(* Logix 5000 project; controller OWF Emulate 5570 rev 30.12; software revision 30.00 *)

TASK MainTask (periodic, rate 1000 ms, priority 1, watchdog 5000 ms) : MainProgram

MODULES
   Local : Emulate 5570 (ICP 2, rev 30.12)
       : vendor 1 type 0 code 15 (ICP 0, rev 1.1, Output RPI 50 ms)
END_MODULES

TYPE UDT_BA :
STRUCT
   AL : BOOL[128];
END_STRUCT
END_TYPE

PROGRAM MainProgram   (* main routine MainRoutine *)
VAR
   OWF_Add_c : DINT;
   OWF_bit : DINT;
   OWF_blk : DINT;
   OWF_i : DINT;
   OWF_Input : DINT[16];
   OWF_InputLen : DINT;
   OWF_InputMaxInd : DINT;
   OWF_j : DINT;
   OWF_Key : DINT[512,17];
   OWF_Result : DINT[17];
   OWF_Ver : DINT;
   SCAN_CYCLE_TIME : DINT;
END_VAR

ROUTINE Application   (* structured text *)
   //Description: initialize the variables.
   
   if S:FS then  (* this is the first, normal scan of the routines in the current program, initialize the program.*)
   	OWF_Ver:=2;  //OWF_Ver means that the version of OWF: 256-256 bits, 384-384 bits, and 512-512 bits. The first number is length of input, the last number is length of output.
                    //If OWF_Ver means that the version of Hash, then three versions are: 256-128 bits, 384-160 bits and 512-256 bits.
   	If OWF_Ver=0 then
   		OWF_InputLen:=255;  //bits of input.
   		OWF_InputMaxInd:=8;  //maximum index for dints which store the bits of input.
   		for OWF_i:=0 to OWF_InputMaxInd-1 by 1 Do
   			//OWF_Input[OWF_i]:= 65535;   //Half of the selection factors are 1.
   			OWF_Input[OWF_i]:= -1;    //All the selection factors are 1.
   		end_for;
   	end_if;
   
   
   	If OWF_Ver=1 then
   		OWF_InputLen:= 383;
   		OWF_InputMaxInd:=12;  //maximum index for array.
   		for OWF_i:=0 to OWF_InputMaxInd-1 by 1 Do
   			//OWF_Input[OWF_i]:= 65535;     //Half of the selection factors are 1.
   			OWF_Input[OWF_i]:= -1;   //All the selection factors are 1.
   		end_for;
   	end_if;
   
   
   	If OWF_Ver=2 then
   		OWF_InputLen:= 511;
   		OWF_InputMaxInd:=16;  //maximum index for array.
   		for OWF_i:=0 to OWF_InputMaxInd-1 by 1 Do
   			//OWF_Input[OWF_i]:= 65535;     //Half of the selection factors are 1.
   			OWF_Input[OWF_i]:= -1;   //All the selection factors are 1.
   		end_for;
   	end_if;
   
   end_if;
   
   
   
   
   
END_ROUTINE

ROUTINE MainRoutine   (* ladder *)
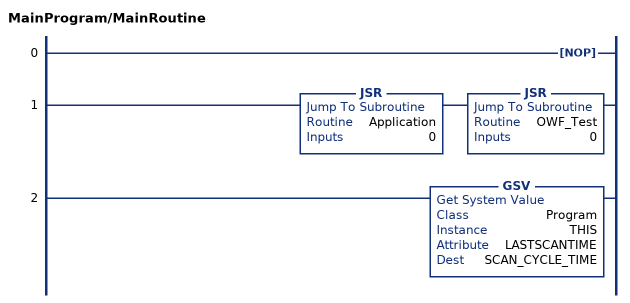
   0: NOP();
   1: JSR(Application,0)JSR(OWF_Test,0);
   2: GSV(Program,THIS,LASTSCANTIME,SCAN_CYCLE_TIME);
END_ROUTINE

ROUTINE Original_OWF   (* structured text *)
   
   //implement One Way Function (OWF) based on subset Sum.
   //input: choice factor OWF_Input[], array OWF_Key[][].
   //output: OWF_Result[]
   
   (*
   	for OWF_i:=0 to OWF_InputMaxInd by 1 Do
   		OWF_Result[OWF_i]:= 0;  //Initialize the OWF_Result[].
   	end_for;
   *)
   
   
   OWF_bit:=0;   // bit index
   OWF_blk:=0;   // block index
   
   JSR(OWF_Init);
   
   	//compute subset sum.
   	for OWF_i:=0 to OWF_InputLen by 1 do
   		If OWF_bit = 32 then
   			OWF_bit:=0;
   			OWF_blk:=OWF_blk+1;
   		end_if;
   		OWF_Add_c:=0;
   		if OWF_Input[OWF_blk].[OWF_bit] then
   			for OWF_j:=0 to OWF_InputMaxInd-1 by 1 Do
   				OWF_Result[OWF_j]:=OWF_Result[OWF_j] + OWF_Key[OWF_i,OWF_j] + OWF_Add_c;    //compute the result of subset sum.
   				OWF_Add_c.0:= OWF_Result[OWF_j].31;
   				OWF_Result[OWF_j].31:=0;
   			end_for;
   			OWF_Result[OWF_j]:=OWF_Result[OWF_j] + OWF_Key[OWF_i,OWF_j] + OWF_Add_c;
   		end_if;
   		OWF_bit:=OWF_bit + 1;
   	end_for;
   
   If OWF_Ver=0 Then
   	OWF_Result[OWF_InputMaxInd]:=OWF_Result[OWF_InputMaxInd] and 16#FF; //clear high bit
   End_If;
   
   If OWF_Ver=1 Then
   	OWF_Result[OWF_InputMaxInd]:=OWF_Result[OWF_InputMaxInd] and 16#FFF; //clear high bit
   End_If;
   
   If OWF_Ver = 2 Then
   	OWF_Result[OWF_InputMaxInd]:=OWF_Result[OWF_InputMaxInd] and 16#FFFF; //clear high bit
   End_If;
END_ROUTINE

ROUTINE OWF_Init   (* structured text *)
   If OWF_Ver >= 0 Then
   	OWF_Key[0,0]:=1227121054;
   	OWF_Key[0,1]:=202649963;
   	OWF_Key[0,2]:=1031163235;
   	OWF_Key[0,3]:=558332383;
   	OWF_Key[0,4]:=758449748;
   	OWF_Key[0,5]:=439100062;
   	OWF_Key[0,6]:=1763017217;
   	OWF_Key[0,7]:=741113131;
   	OWF_Key[0,8]:=1652892808;
   	OWF_Key[1,0]:=1354606577;
   	OWF_Key[1,1]:=1085346626;
   	OWF_Key[1,2]:=1684734244;
   	OWF_Key[1,3]:=1525280682;
   	OWF_Key[1,4]:=581896247;
   	OWF_Key[1,5]:=1418880834;
   	OWF_Key[1,6]:=1348359995;
   	OWF_Key[1,7]:=1446005479;
   	OWF_Key[1,8]:=332839494;
   	OWF_Key[2,0]:=2095017041;
   	OWF_Key[2,1]:=1217317816;
   	OWF_Key[2,2]:=648181522;
   	OWF_Key[2,3]:=178964298;
   	OWF_Key[2,4]:=463461758;
   	OWF_Key[2,5]:=346394231;
   	OWF_Key[2,6]:=1486999699;
   	OWF_Key[2,7]:=1770617031;
   	OWF_Key[2,8]:=362139479;
   	OWF_Key[3,0]:=256347809;
   	OWF_Key[3,1]:=1312207174;
   	OWF_Key[3,2]:=843085075;
   	OWF_Key[3,3]:=1139982972;
   	OWF_Key[3,4]:=662387156;
   	OWF_Key[3,5]:=1025052915;
   	OWF_Key[3,6]:=1908648583;
   	OWF_Key[3,7]:=1963224943;
   	OWF_Key[3,8]:=1427256681;
   	OWF_Key[4,0]:=1972101745;
   	OWF_Key[4,1]:=1002975333;
   	OWF_Key[4,2]:=1871427740;
   	OWF_Key[4,3]:=1318551426;
   	OWF_Key[4,4]:=1364597906;
   	OWF_Key[4,5]:=1294123204;
   	OWF_Key[4,6]:=2125414218;
   	OWF_Key[4,7]:=1926341024;
   	OWF_Key[4,8]:=460259043;
   	OWF_Key[5,0]:=1524399156;
   	OWF_Key[5,1]:=2011514619;
   	OWF_Key[5,2]:=2069350563;
   	OWF_Key[5,3]:=279858814;
   	OWF_Key[5,4]:=810485067;
   	OWF_Key[5,5]:=73617388;
   	OWF_Key[5,6]:=687884215;
   	OWF_Key[5,7]:=1340310677;
   	OWF_Key[5,8]:=431345285;
   	OWF_Key[6,0]:=1066476071;
   	OWF_Key[6,1]:=550806088;
   	OWF_Key[6,2]:=756174308;
   	OWF_Key[6,3]:=574071763;
   	OWF_Key[6,4]:=409094206;
   	OWF_Key[6,5]:=1665642823;
   	OWF_Key[6,6]:=1813040245;
   	OWF_Key[6,7]:=215573695;
   	OWF_Key[6,8]:=525097691;
   	OWF_Key[7,0]:=1934399231;
   	OWF_Key[7,1]:=1553053230;
   	OWF_Key[7,2]:=144946822;
   	OWF_Key[7,3]:=2140599730;
   	OWF_Key[7,4]:=1889193085;
   	OWF_Key[7,5]:=2054644962;
   	OWF_Key[7,6]:=826013297;
   	OWF_Key[7,7]:=556817065;
   	OWF_Key[7,8]:=33718400;
   	OWF_Key[8,0]:=899651387;
   	OWF_Key[8,1]:=1251867014;
   	OWF_Key[8,2]:=959094800;
   	OWF_Key[8,3]:=194574689;
   	OWF_Key[8,4]:=1642465144;
   	OWF_Key[8,5]:=1096334976;
   	OWF_Key[8,6]:=931056050;
   	OWF_Key[8,7]:=405780298;
   	OWF_Key[8,8]:=1355752490;
   	OWF_Key[9,0]:=1528579024;
   	OWF_Key[9,1]:=1525333419;
   	OWF_Key[9,2]:=1348534735;
   	OWF_Key[9,3]:=111603084;
   	OWF_Key[9,4]:=1832745100;
   	OWF_Key[9,5]:=642195240;
   	OWF_Key[9,6]:=966181946;
   	OWF_Key[9,7]:=880029259;
   	OWF_Key[9,8]:=1162642342;
   	OWF_Key[10,0]:=359569674;
   	OWF_Key[10,1]:=1980700574;
   	OWF_Key[10,2]:=1293914236;
   	OWF_Key[10,3]:=954723255;
   	OWF_Key[10,4]:=1377909373;
   	OWF_Key[10,5]:=223244700;
   	OWF_Key[10,6]:=1984808221;
   	OWF_Key[10,7]:=1498924409;
   	OWF_Key[10,8]:=29167191;
   	OWF_Key[11,0]:=623116396;
   	OWF_Key[11,1]:=256225512;
   	OWF_Key[11,2]:=1328608936;
   	OWF_Key[11,3]:=725706243;
   	OWF_Key[11,4]:=791017754;
   	OWF_Key[11,5]:=1341758946;
   	OWF_Key[11,6]:=1113167772;
   	OWF_Key[11,7]:=639937104;
   	OWF_Key[11,8]:=436330960;
   	OWF_Key[12,0]:=1329424307;
   	OWF_Key[12,1]:=101924380;
   	OWF_Key[12,2]:=1635207076;
   	OWF_Key[12,3]:=1264309098;
   	OWF_Key[12,4]:=1613321141;
   	OWF_Key[12,5]:=1843793655;
   	OWF_Key[12,6]:=1519128380;
   	OWF_Key[12,7]:=1637695475;
   	OWF_Key[12,8]:=1595160782;
   	OWF_Key[13,0]:=475438733;
   	OWF_Key[13,1]:=914493831;
   	OWF_Key[13,2]:=239185193;
   	OWF_Key[13,3]:=7070920;
   	OWF_Key[13,4]:=1909091689;
   	OWF_Key[13,5]:=818931882;
   	OWF_Key[13,6]:=167044628;
   	OWF_Key[13,7]:=1264941904;
   	OWF_Key[13,8]:=949875305;
   	OWF_Key[14,0]:=1115356298;
   	OWF_Key[14,1]:=338497818;
   	OWF_Key[14,2]:=180024891;
   	OWF_Key[14,3]:=844456349;
   	OWF_Key[14,4]:=1506829383;
   	OWF_Key[14,5]:=94052327;
   	OWF_Key[14,6]:=1993991460;
   	OWF_Key[14,7]:=23038222;
   	OWF_Key[14,8]:=87146691;
   	OWF_Key[15,0]:=326487164;
   	OWF_Key[15,1]:=516484364;
   	OWF_Key[15,2]:=1296941749;
   	OWF_Key[15,3]:=811092697;
   	OWF_Key[15,4]:=538927605;
   	OWF_Key[15,5]:=659414599;
   	OWF_Key[15,6]:=759387250;
   	OWF_Key[15,7]:=589772068;
   	OWF_Key[15,8]:=514624038;
   	OWF_Key[16,0]:=1091875462;
   	OWF_Key[16,1]:=461268148;
   	OWF_Key[16,2]:=1603288957;
   	OWF_Key[16,3]:=626416433;
   	OWF_Key[16,4]:=654301897;
   	OWF_Key[16,5]:=1861165437;
   	OWF_Key[16,6]:=710648683;
   	OWF_Key[16,7]:=706991177;
   	OWF_Key[16,8]:=2023521577;
   	OWF_Key[17,0]:=1533914360;
   	OWF_Key[17,1]:=2033382504;
   	OWF_Key[17,2]:=1913483458;
   	OWF_Key[17,3]:=1068320764;
   	OWF_Key[17,4]:=1873217994;
   	OWF_Key[17,5]:=462057421;
   	OWF_Key[17,6]:=434206996;
   	OWF_Key[17,7]:=967662215;
   	OWF_Key[17,8]:=1066362328;
   	OWF_Key[18,0]:=1233616361;
   	OWF_Key[18,1]:=1376108010;
   	OWF_Key[18,2]:=151681671;
   	OWF_Key[18,3]:=1118724616;
   	OWF_Key[18,4]:=870582805;
   	OWF_Key[18,5]:=838422454;
   	OWF_Key[18,6]:=958525863;
   	OWF_Key[18,7]:=884926077;
   	OWF_Key[18,8]:=1110871443;
   	OWF_Key[19,0]:=1105934356;
   	OWF_Key[19,1]:=664442467;
   	OWF_Key[19,2]:=903233013;
   	OWF_Key[19,3]:=987099294;
   	OWF_Key[19,4]:=737604300;
   	OWF_Key[19,5]:=1759631091;
   	OWF_Key[19,6]:=1580233890;
   	OWF_Key[19,7]:=1669577827;
   	OWF_Key[19,8]:=91657386;
   	OWF_Key[20,0]:=360120849;
   	OWF_Key[20,1]:=1832314473;
   	OWF_Key[20,2]:=2086185527;
   	OWF_Key[20,3]:=1076864314;
   	OWF_Key[20,4]:=1498905358;
   	OWF_Key[20,5]:=900988985;
   	OWF_Key[20,6]:=1478986721;
   	OWF_Key[20,7]:=1681057774;
   	OWF_Key[20,8]:=562389748;
   	OWF_Key[21,0]:=368575225;
   	OWF_Key[21,1]:=2040057957;
   	OWF_Key[21,2]:=1772443406;
   	OWF_Key[21,3]:=358038348;
   	OWF_Key[21,4]:=1880468616;
   	OWF_Key[21,5]:=1275762442;
   	OWF_Key[21,6]:=240738790;
   	OWF_Key[21,7]:=1742748974;
   	OWF_Key[21,8]:=1288995313;
   	OWF_Key[22,0]:=2102585710;
   	OWF_Key[22,1]:=1254850839;
   	OWF_Key[22,2]:=1750685415;
   	OWF_Key[22,3]:=407311703;
   	OWF_Key[22,4]:=1927455536;
   	OWF_Key[22,5]:=734780728;
   	OWF_Key[22,6]:=1963803180;
   	OWF_Key[22,7]:=24276587;
   	OWF_Key[22,8]:=305836334;
   	OWF_Key[23,0]:=1060880211;
   	OWF_Key[23,1]:=321236053;
   	OWF_Key[23,2]:=1978313959;
   	OWF_Key[23,3]:=280999634;
   	OWF_Key[23,4]:=811422929;
   	OWF_Key[23,5]:=1151495141;
   	OWF_Key[23,6]:=684998164;
   	OWF_Key[23,7]:=1774640068;
   	OWF_Key[23,8]:=1081430675;
   	OWF_Key[24,0]:=1100474918;
   	OWF_Key[24,1]:=604700422;
   	OWF_Key[24,2]:=1689758319;
   	OWF_Key[24,3]:=215570041;
   	OWF_Key[24,4]:=1701438018;
   	OWF_Key[24,5]:=1754755041;
   	OWF_Key[24,6]:=7425442;
   	OWF_Key[24,7]:=918208170;
   	OWF_Key[24,8]:=1719377360;
   	OWF_Key[25,0]:=1547355790;
   	OWF_Key[25,1]:=1403608030;
   	OWF_Key[25,2]:=1499880269;
   	OWF_Key[25,3]:=317100104;
   	OWF_Key[25,4]:=1905628845;
   	OWF_Key[25,5]:=1066486402;
   	OWF_Key[25,6]:=756239231;
   	OWF_Key[25,7]:=459531339;
   	OWF_Key[25,8]:=1346452392;
   	OWF_Key[26,0]:=168483711;
   	OWF_Key[26,1]:=1800574949;
   	OWF_Key[26,2]:=1200797705;
   	OWF_Key[26,3]:=14565181;
   	OWF_Key[26,4]:=228173521;
   	OWF_Key[26,5]:=1764496443;
   	OWF_Key[26,6]:=504637489;
   	OWF_Key[26,7]:=1780840621;
   	OWF_Key[26,8]:=1379082303;
   	OWF_Key[27,0]:=54123181;
   	OWF_Key[27,1]:=622944351;
   	OWF_Key[27,2]:=2100500392;
   	OWF_Key[27,3]:=1775742704;
   	OWF_Key[27,4]:=143633756;
   	OWF_Key[27,5]:=1536231566;
   	OWF_Key[27,6]:=1440183257;
   	OWF_Key[27,7]:=2114239512;
   	OWF_Key[27,8]:=53396177;
   	OWF_Key[28,0]:=2134211248;
   	OWF_Key[28,1]:=1985332782;
   	OWF_Key[28,2]:=660997500;
   	OWF_Key[28,3]:=1607311701;
   	OWF_Key[28,4]:=1401991464;
   	OWF_Key[28,5]:=891355717;
   	OWF_Key[28,6]:=1475041716;
   	OWF_Key[28,7]:=258011330;
   	OWF_Key[28,8]:=2098653906;
   	OWF_Key[29,0]:=1790937980;
   	OWF_Key[29,1]:=592851196;
   	OWF_Key[29,2]:=1910540181;
   	OWF_Key[29,3]:=664243004;
   	OWF_Key[29,4]:=360474841;
   	OWF_Key[29,5]:=1110300911;
   	OWF_Key[29,6]:=1039400747;
   	OWF_Key[29,7]:=404077093;
   	OWF_Key[29,8]:=1245988018;
   	OWF_Key[30,0]:=82206939;
   	OWF_Key[30,1]:=2105921183;
   	OWF_Key[30,2]:=586971854;
   	OWF_Key[30,3]:=1765305131;
   	OWF_Key[30,4]:=1096912113;
   	OWF_Key[30,5]:=1614673633;
   	OWF_Key[30,6]:=899093717;
   	OWF_Key[30,7]:=476264675;
   	OWF_Key[30,8]:=958189495;
   	OWF_Key[31,0]:=1427661975;
   	OWF_Key[31,1]:=2139629653;
   	OWF_Key[31,2]:=922325329;
   	OWF_Key[31,3]:=139475207;
   	OWF_Key[31,4]:=864976279;
   	OWF_Key[31,5]:=115584651;
   	OWF_Key[31,6]:=1609825306;
   	OWF_Key[31,7]:=1667460585;
   	OWF_Key[31,8]:=1143913594;
   	OWF_Key[32,0]:=1568245993;
   	OWF_Key[32,1]:=1049047354;
   	OWF_Key[32,2]:=959206126;
   	OWF_Key[32,3]:=1741588568;
   	OWF_Key[32,4]:=1470670599;
   	OWF_Key[32,5]:=1694909057;
   	OWF_Key[32,6]:=235889822;
   	OWF_Key[32,7]:=3720639;
   	OWF_Key[32,8]:=125832420;
   	OWF_Key[33,0]:=648198321;
   	OWF_Key[33,1]:=1530796919;
   	OWF_Key[33,2]:=1793974282;
   	OWF_Key[33,3]:=1628769796;
   	OWF_Key[33,4]:=1884925188;
   	OWF_Key[33,5]:=401471910;
   	OWF_Key[33,6]:=928541632;
   	OWF_Key[33,7]:=881114955;
   	OWF_Key[33,8]:=533672300;
   	OWF_Key[34,0]:=1343614706;
   	OWF_Key[34,1]:=1565280378;
   	OWF_Key[34,2]:=1934951256;
   	OWF_Key[34,3]:=1283078343;
   	OWF_Key[34,4]:=516108734;
   	OWF_Key[34,5]:=1739049325;
   	OWF_Key[34,6]:=1170335756;
   	OWF_Key[34,7]:=913104818;
   	OWF_Key[34,8]:=86599362;
   	OWF_Key[35,0]:=1657291640;
   	OWF_Key[35,1]:=1813687561;
   	OWF_Key[35,2]:=1076706992;
   	OWF_Key[35,3]:=1082055811;
   	OWF_Key[35,4]:=858507228;
   	OWF_Key[35,5]:=566669145;
   	OWF_Key[35,6]:=235309761;
   	OWF_Key[35,7]:=890380619;
   	OWF_Key[35,8]:=1422472402;
   	OWF_Key[36,0]:=1446507793;
   	OWF_Key[36,1]:=1328829415;
   	OWF_Key[36,2]:=1380176807;
   	OWF_Key[36,3]:=1633730348;
   	OWF_Key[36,4]:=745778942;
   	OWF_Key[36,5]:=1055032828;
   	OWF_Key[36,6]:=1520091153;
   	OWF_Key[36,7]:=1535317210;
   	OWF_Key[36,8]:=1044560664;
   	OWF_Key[37,0]:=604110439;
   	OWF_Key[37,1]:=26486716;
   	OWF_Key[37,2]:=2049306560;
   	OWF_Key[37,3]:=1798262270;
   	OWF_Key[37,4]:=1200653570;
   	OWF_Key[37,5]:=249378793;
   	OWF_Key[37,6]:=1132886992;
   	OWF_Key[37,7]:=1600976401;
   	OWF_Key[37,8]:=819015577;
   	OWF_Key[38,0]:=76994523;
   	OWF_Key[38,1]:=491360675;
   	OWF_Key[38,2]:=576400950;
   	OWF_Key[38,3]:=1590171180;
   	OWF_Key[38,4]:=115692894;
   	OWF_Key[38,5]:=739418327;
   	OWF_Key[38,6]:=1054282547;
   	OWF_Key[38,7]:=584979767;
   	OWF_Key[38,8]:=1253169315;
   	OWF_Key[39,0]:=411932280;
   	OWF_Key[39,1]:=272616828;
   	OWF_Key[39,2]:=239495733;
   	OWF_Key[39,3]:=1888586440;
   	OWF_Key[39,4]:=831515848;
   	OWF_Key[39,5]:=1268168776;
   	OWF_Key[39,6]:=1600339397;
   	OWF_Key[39,7]:=978596994;
   	OWF_Key[39,8]:=53521075;
   	OWF_Key[40,0]:=782007485;
   	OWF_Key[40,1]:=547761025;
   	OWF_Key[40,2]:=1788398174;
   	OWF_Key[40,3]:=1858267849;
   	OWF_Key[40,4]:=86296681;
   	OWF_Key[40,5]:=478881018;
   	OWF_Key[40,6]:=231000794;
   	OWF_Key[40,7]:=453896809;
   	OWF_Key[40,8]:=1637170327;
   	OWF_Key[41,0]:=673014602;
   	OWF_Key[41,1]:=720938492;
   	OWF_Key[41,2]:=749952923;
   	OWF_Key[41,3]:=960648251;
   	OWF_Key[41,4]:=576682832;
   	OWF_Key[41,5]:=1888044580;
   	OWF_Key[41,6]:=1258761492;
   	OWF_Key[41,7]:=1081332593;
   	OWF_Key[41,8]:=1992300120;
   	OWF_Key[42,0]:=1132458609;
   	OWF_Key[42,1]:=548052059;
   	OWF_Key[42,2]:=1506585657;
   	OWF_Key[42,3]:=1131409825;
   	OWF_Key[42,4]:=859232979;
   	OWF_Key[42,5]:=1613011416;
   	OWF_Key[42,6]:=985832894;
   	OWF_Key[42,7]:=965782405;
   	OWF_Key[42,8]:=1483700964;
   	OWF_Key[43,0]:=1009032951;
   	OWF_Key[43,1]:=1777279179;
   	OWF_Key[43,2]:=739680041;
   	OWF_Key[43,3]:=443997529;
   	OWF_Key[43,4]:=824225282;
   	OWF_Key[43,5]:=32764525;
   	OWF_Key[43,6]:=378580490;
   	OWF_Key[43,7]:=680945380;
   	OWF_Key[43,8]:=369690021;
   	OWF_Key[44,0]:=1640626484;
   	OWF_Key[44,1]:=1561378686;
   	OWF_Key[44,2]:=1095897085;
   	OWF_Key[44,3]:=1195403520;
   	OWF_Key[44,4]:=325645116;
   	OWF_Key[44,5]:=1091014514;
   	OWF_Key[44,6]:=541535695;
   	OWF_Key[44,7]:=286402630;
   	OWF_Key[44,8]:=1102658970;
   	OWF_Key[45,0]:=1002827150;
   	OWF_Key[45,1]:=352381150;
   	OWF_Key[45,2]:=1335011513;
   	OWF_Key[45,3]:=245363487;
   	OWF_Key[45,4]:=1029590752;
   	OWF_Key[45,5]:=856290625;
   	OWF_Key[45,6]:=802555697;
   	OWF_Key[45,7]:=329424908;
   	OWF_Key[45,8]:=2104840495;
   	OWF_Key[46,0]:=1665300904;
   	OWF_Key[46,1]:=209108703;
   	OWF_Key[46,2]:=1779396682;
   	OWF_Key[46,3]:=1256656350;
   	OWF_Key[46,4]:=191441463;
   	OWF_Key[46,5]:=1797343127;
   	OWF_Key[46,6]:=2055633172;
   	OWF_Key[46,7]:=584162859;
   	OWF_Key[46,8]:=39760195;
   	OWF_Key[47,0]:=41354911;
   	OWF_Key[47,1]:=1199557050;
   	OWF_Key[47,2]:=1765662309;
   	OWF_Key[47,3]:=551500113;
   	OWF_Key[47,4]:=1511913983;
   	OWF_Key[47,5]:=2018316238;
   	OWF_Key[47,6]:=1666070399;
   	OWF_Key[47,7]:=1342412915;
   	OWF_Key[47,8]:=842109359;
   	OWF_Key[48,0]:=705031084;
   	OWF_Key[48,1]:=108181531;
   	OWF_Key[48,2]:=211069878;
   	OWF_Key[48,3]:=1128443167;
   	OWF_Key[48,4]:=664585396;
   	OWF_Key[48,5]:=1761822658;
   	OWF_Key[48,6]:=142165939;
   	OWF_Key[48,7]:=535769991;
   	OWF_Key[48,8]:=239150875;
   	OWF_Key[49,0]:=140746729;
   	OWF_Key[49,1]:=146417569;
   	OWF_Key[49,2]:=1111962022;
   	OWF_Key[49,3]:=1720219764;
   	OWF_Key[49,4]:=1351513412;
   	OWF_Key[49,5]:=1975372593;
   	OWF_Key[49,6]:=1521231143;
   	OWF_Key[49,7]:=592752896;
   	OWF_Key[49,8]:=1716537172;
   	OWF_Key[50,0]:=1289831067;
   	OWF_Key[50,1]:=556791851;
   	OWF_Key[50,2]:=1601279844;
   	OWF_Key[50,3]:=1113008242;
   	OWF_Key[50,4]:=257492968;
   	OWF_Key[50,5]:=448491471;
   	OWF_Key[50,6]:=1348139853;
   	OWF_Key[50,7]:=1265875548;
   	OWF_Key[50,8]:=1112480858;
   	OWF_Key[51,0]:=958741303;
   	OWF_Key[51,1]:=625050139;
   	OWF_Key[51,2]:=1907318927;
   	OWF_Key[51,3]:=1790227796;
   	OWF_Key[51,4]:=982526424;
   	OWF_Key[51,5]:=403675080;
   	OWF_Key[51,6]:=1159748236;
   	OWF_Key[51,7]:=1367875897;
   	OWF_Key[51,8]:=232916365;
   	OWF_Key[52,0]:=1517162145;
   	OWF_Key[52,1]:=2088172931;
   	OWF_Key[52,2]:=962493317;
   	OWF_Key[52,3]:=1067933972;
   	OWF_Key[52,4]:=1327199334;
   	OWF_Key[52,5]:=610006435;
   	OWF_Key[52,6]:=2109925092;
   	OWF_Key[52,7]:=1068942317;
   	OWF_Key[52,8]:=173113135;
   	OWF_Key[53,0]:=1278524224;
   	OWF_Key[53,1]:=1252167227;
   	OWF_Key[53,2]:=1127816425;
   	OWF_Key[53,3]:=145099354;
   	OWF_Key[53,4]:=1487037740;
   	OWF_Key[53,5]:=1734599138;
   	OWF_Key[53,6]:=141607975;
   	OWF_Key[53,7]:=1228460997;
   	OWF_Key[53,8]:=1261511827;
   	OWF_Key[54,0]:=991465721;
   	OWF_Key[54,1]:=1620985555;
   	OWF_Key[54,2]:=1976927632;
   	OWF_Key[54,3]:=1882638804;
   	OWF_Key[54,4]:=223756234;
   	OWF_Key[54,5]:=882310812;
   	OWF_Key[54,6]:=1952374609;
   	OWF_Key[54,7]:=1588702672;
   	OWF_Key[54,8]:=672111005;
   	OWF_Key[55,0]:=173274277;
   	OWF_Key[55,1]:=1842190662;
   	OWF_Key[55,2]:=45228216;
   	OWF_Key[55,3]:=1986844369;
   	OWF_Key[55,4]:=2024468617;
   	OWF_Key[55,5]:=1745946897;
   	OWF_Key[55,6]:=1215380589;
   	OWF_Key[55,7]:=200791282;
   	OWF_Key[55,8]:=1300581522;
   	OWF_Key[56,0]:=1834029440;
   	OWF_Key[56,1]:=1363563541;
   	OWF_Key[56,2]:=535408957;
   	OWF_Key[56,3]:=469857245;
   	OWF_Key[56,4]:=675815278;
   	OWF_Key[56,5]:=1278408349;
   	OWF_Key[56,6]:=933515210;
   	OWF_Key[56,7]:=1316646286;
   	OWF_Key[56,8]:=373047480;
   	OWF_Key[57,0]:=1016144636;
   	OWF_Key[57,1]:=1779677369;
   	OWF_Key[57,2]:=58728151;
   	OWF_Key[57,3]:=1358234411;
   	OWF_Key[57,4]:=1834858672;
   	OWF_Key[57,5]:=1406013272;
   	OWF_Key[57,6]:=1423437632;
   	OWF_Key[57,7]:=1421089637;
   	OWF_Key[57,8]:=1985019890;
   	OWF_Key[58,0]:=1580033881;
   	OWF_Key[58,1]:=457883305;
   	OWF_Key[58,2]:=470943474;
   	OWF_Key[58,3]:=923583801;
   	OWF_Key[58,4]:=1769010706;
   	OWF_Key[58,5]:=1375307187;
   	OWF_Key[58,6]:=363536141;
   	OWF_Key[58,7]:=1121047259;
   	OWF_Key[58,8]:=1061644749;
   	OWF_Key[59,0]:=1475052699;
   	OWF_Key[59,1]:=1021043562;
   	OWF_Key[59,2]:=207530477;
   	OWF_Key[59,3]:=1655456205;
   	OWF_Key[59,4]:=851724661;
   	OWF_Key[59,5]:=1116609908;
   	OWF_Key[59,6]:=1200895844;
   	OWF_Key[59,7]:=2108312592;
   	OWF_Key[59,8]:=1849271216;
   	OWF_Key[60,0]:=470886666;
   	OWF_Key[60,1]:=430952018;
   	OWF_Key[60,2]:=1420232976;
   	OWF_Key[60,3]:=526556583;
   	OWF_Key[60,4]:=1340856141;
   	OWF_Key[60,5]:=682182388;
   	OWF_Key[60,6]:=1657105479;
   	OWF_Key[60,7]:=826355643;
   	OWF_Key[60,8]:=1023121452;
   	OWF_Key[61,0]:=1850440524;
   	OWF_Key[61,1]:=314641402;
   	OWF_Key[61,2]:=340220969;
   	OWF_Key[61,3]:=1494492295;
   	OWF_Key[61,4]:=402187581;
   	OWF_Key[61,5]:=877825514;
   	OWF_Key[61,6]:=119246503;
   	OWF_Key[61,7]:=346949548;
   	OWF_Key[61,8]:=490871209;
   	OWF_Key[62,0]:=2123319554;
   	OWF_Key[62,1]:=1040649935;
   	OWF_Key[62,2]:=2058114642;
   	OWF_Key[62,3]:=1246595551;
   	OWF_Key[62,4]:=1344918190;
   	OWF_Key[62,5]:=1749844790;
   	OWF_Key[62,6]:=70180448;
   	OWF_Key[62,7]:=1492229206;
   	OWF_Key[62,8]:=1974255998;
   	OWF_Key[63,0]:=826345708;
   	OWF_Key[63,1]:=569432486;
   	OWF_Key[63,2]:=1662176022;
   	OWF_Key[63,3]:=1069949292;
   	OWF_Key[63,4]:=3045329;
   	OWF_Key[63,5]:=1948384876;
   	OWF_Key[63,6]:=2132761985;
   	OWF_Key[63,7]:=1556848512;
   	OWF_Key[63,8]:=773814376;
   	OWF_Key[64,0]:=1967105076;
   	OWF_Key[64,1]:=718865195;
   	OWF_Key[64,2]:=843916660;
   	OWF_Key[64,3]:=594129844;
   	OWF_Key[64,4]:=1571287676;
   	OWF_Key[64,5]:=1651982779;
   	OWF_Key[64,6]:=155599888;
   	OWF_Key[64,7]:=1337181185;
   	OWF_Key[64,8]:=1969333902;
   	OWF_Key[65,0]:=375598944;
   	OWF_Key[65,1]:=1899047934;
   	OWF_Key[65,2]:=2014896421;
   	OWF_Key[65,3]:=29097043;
   	OWF_Key[65,4]:=217403893;
   	OWF_Key[65,5]:=463855642;
   	OWF_Key[65,6]:=1482864454;
   	OWF_Key[65,7]:=956236890;
   	OWF_Key[65,8]:=518322261;
   	OWF_Key[66,0]:=497089837;
   	OWF_Key[66,1]:=1705294572;
   	OWF_Key[66,2]:=1369872479;
   	OWF_Key[66,3]:=1950228985;
   	OWF_Key[66,4]:=822587228;
   	OWF_Key[66,5]:=1306639444;
   	OWF_Key[66,6]:=901234665;
   	OWF_Key[66,7]:=1370427942;
   	OWF_Key[66,8]:=279387629;
   	OWF_Key[67,0]:=160995784;
   	OWF_Key[67,1]:=533581559;
   	OWF_Key[67,2]:=1980127655;
   	OWF_Key[67,3]:=1562262632;
   	OWF_Key[67,4]:=1117184000;
   	OWF_Key[67,5]:=1662051811;
   	OWF_Key[67,6]:=883414987;
   	OWF_Key[67,7]:=707506599;
   	OWF_Key[67,8]:=1614769155;
   	OWF_Key[68,0]:=821129193;
   	OWF_Key[68,1]:=1231377393;
   	OWF_Key[68,2]:=209468532;
   	OWF_Key[68,3]:=48572430;
   	OWF_Key[68,4]:=914969677;
   	OWF_Key[68,5]:=1107553125;
   	OWF_Key[68,6]:=1203724242;
   	OWF_Key[68,7]:=802136307;
   	OWF_Key[68,8]:=2132413638;
   	OWF_Key[69,0]:=1753436816;
   	OWF_Key[69,1]:=1515658151;
   	OWF_Key[69,2]:=1696060662;
   	OWF_Key[69,3]:=1440580301;
   	OWF_Key[69,4]:=1232973813;
   	OWF_Key[69,5]:=622697960;
   	OWF_Key[69,6]:=1033056322;
   	OWF_Key[69,7]:=1236071203;
   	OWF_Key[69,8]:=1123543335;
   	OWF_Key[70,0]:=1313474539;
   	OWF_Key[70,1]:=25955154;
   	OWF_Key[70,2]:=1500583878;
   	OWF_Key[70,3]:=2108697879;
   	OWF_Key[70,4]:=82386448;
   	OWF_Key[70,5]:=872426545;
   	OWF_Key[70,6]:=688921535;
   	OWF_Key[70,7]:=222876749;
   	OWF_Key[70,8]:=594319329;
   	OWF_Key[71,0]:=699509228;
   	OWF_Key[71,1]:=371806453;
   	OWF_Key[71,2]:=469265036;
   	OWF_Key[71,3]:=1179216536;
   	OWF_Key[71,4]:=1525572509;
   	OWF_Key[71,5]:=876866338;
   	OWF_Key[71,6]:=2107468087;
   	OWF_Key[71,7]:=580688836;
   	OWF_Key[71,8]:=922828615;
   	OWF_Key[72,0]:=1551486097;
   	OWF_Key[72,1]:=1862819700;
   	OWF_Key[72,2]:=1601215303;
   	OWF_Key[72,3]:=847797762;
   	OWF_Key[72,4]:=1142119955;
   	OWF_Key[72,5]:=1730944373;
   	OWF_Key[72,6]:=761903716;
   	OWF_Key[72,7]:=476549925;
   	OWF_Key[72,8]:=742414564;
   	OWF_Key[73,0]:=1983411600;
   	OWF_Key[73,1]:=452261303;
   	OWF_Key[73,2]:=597231909;
   	OWF_Key[73,3]:=1125992219;
   	OWF_Key[73,4]:=1912687650;
   	OWF_Key[73,5]:=1727260970;
   	OWF_Key[73,6]:=316209247;
   	OWF_Key[73,7]:=1460211977;
   	OWF_Key[73,8]:=1473283512;
   	OWF_Key[74,0]:=874539113;
   	OWF_Key[74,1]:=1814062959;
   	OWF_Key[74,2]:=1693389721;
   	OWF_Key[74,3]:=1072346191;
   	OWF_Key[74,4]:=2053594629;
   	OWF_Key[74,5]:=680531052;
   	OWF_Key[74,6]:=33202566;
   	OWF_Key[74,7]:=1278556457;
   	OWF_Key[74,8]:=966110963;
   	OWF_Key[75,0]:=1047105521;
   	OWF_Key[75,1]:=170050367;
   	OWF_Key[75,2]:=1921783554;
   	OWF_Key[75,3]:=1702134946;
   	OWF_Key[75,4]:=1686346929;
   	OWF_Key[75,5]:=1348768913;
   	OWF_Key[75,6]:=1098769006;
   	OWF_Key[75,7]:=539879319;
   	OWF_Key[75,8]:=348285647;
   	OWF_Key[76,0]:=1516077301;
   	OWF_Key[76,1]:=1356603304;
   	OWF_Key[76,2]:=1993796975;
   	OWF_Key[76,3]:=1431371711;
   	OWF_Key[76,4]:=1964847289;
   	OWF_Key[76,5]:=1309605544;
   	OWF_Key[76,6]:=415147319;
   	OWF_Key[76,7]:=2006882414;
   	OWF_Key[76,8]:=1279231381;
   	OWF_Key[77,0]:=983568528;
   	OWF_Key[77,1]:=130542355;
   	OWF_Key[77,2]:=1272223238;
   	OWF_Key[77,3]:=2011646589;
   	OWF_Key[77,4]:=1266917943;
   	OWF_Key[77,5]:=70109226;
   	OWF_Key[77,6]:=2032179276;
   	OWF_Key[77,7]:=1345698146;
   	OWF_Key[77,8]:=600376789;
   	OWF_Key[78,0]:=686782273;
   	OWF_Key[78,1]:=1143168531;
   	OWF_Key[78,2]:=630736712;
   	OWF_Key[78,3]:=1667829760;
   	OWF_Key[78,4]:=174554158;
   	OWF_Key[78,5]:=1100164131;
   	OWF_Key[78,6]:=280229495;
   	OWF_Key[78,7]:=686349585;
   	OWF_Key[78,8]:=1415553179;
   	OWF_Key[79,0]:=534407931;
   	OWF_Key[79,1]:=734849944;
   	OWF_Key[79,2]:=1333166045;
   	OWF_Key[79,3]:=2024933309;
   	OWF_Key[79,4]:=256637645;
   	OWF_Key[79,5]:=1721865403;
   	OWF_Key[79,6]:=2062066624;
   	OWF_Key[79,7]:=1918290307;
   	OWF_Key[79,8]:=161209948;
   	OWF_Key[80,0]:=1600364462;
   	OWF_Key[80,1]:=129587141;
   	OWF_Key[80,2]:=1429637701;
   	OWF_Key[80,3]:=1292734676;
   	OWF_Key[80,4]:=1689565378;
   	OWF_Key[80,5]:=1485424925;
   	OWF_Key[80,6]:=1957791753;
   	OWF_Key[80,7]:=225897719;
   	OWF_Key[80,8]:=905680692;
   	OWF_Key[81,0]:=914708458;
   	OWF_Key[81,1]:=1366932185;
   	OWF_Key[81,2]:=998034109;
   	OWF_Key[81,3]:=1218728918;
   	OWF_Key[81,4]:=230333278;
   	OWF_Key[81,5]:=1627616151;
   	OWF_Key[81,6]:=1920189999;
   	OWF_Key[81,7]:=1021983029;
   	OWF_Key[81,8]:=1106545101;
   	OWF_Key[82,0]:=1762097210;
   	OWF_Key[82,1]:=1862139904;
   	OWF_Key[82,2]:=1639202737;
   	OWF_Key[82,3]:=216675238;
   	OWF_Key[82,4]:=1751522393;
   	OWF_Key[82,5]:=982581238;
   	OWF_Key[82,6]:=1093927662;
   	OWF_Key[82,7]:=1191499474;
   	OWF_Key[82,8]:=1428392037;
   	OWF_Key[83,0]:=1290270779;
   	OWF_Key[83,1]:=255582270;
   	OWF_Key[83,2]:=1527656360;
   	OWF_Key[83,3]:=1166394851;
   	OWF_Key[83,4]:=1576211303;
   	OWF_Key[83,5]:=1677433256;
   	OWF_Key[83,6]:=955815081;
   	OWF_Key[83,7]:=1281950671;
   	OWF_Key[83,8]:=1302685485;
   	OWF_Key[84,0]:=1700413184;
   	OWF_Key[84,1]:=839422281;
   	OWF_Key[84,2]:=1123646424;
   	OWF_Key[84,3]:=1318151337;
   	OWF_Key[84,4]:=1742102491;
   	OWF_Key[84,5]:=1546205803;
   	OWF_Key[84,6]:=1160246466;
   	OWF_Key[84,7]:=180580323;
   	OWF_Key[84,8]:=1649852129;
   	OWF_Key[85,0]:=1552429261;
   	OWF_Key[85,1]:=1415057071;
   	OWF_Key[85,2]:=36706649;
   	OWF_Key[85,3]:=28255214;
   	OWF_Key[85,4]:=1722553546;
   	OWF_Key[85,5]:=1745077298;
   	OWF_Key[85,6]:=1107749020;
   	OWF_Key[85,7]:=714530504;
   	OWF_Key[85,8]:=1396093169;
   	OWF_Key[86,0]:=532511322;
   	OWF_Key[86,1]:=493048671;
   	OWF_Key[86,2]:=496742733;
   	OWF_Key[86,3]:=1119913924;
   	OWF_Key[86,4]:=337190732;
   	OWF_Key[86,5]:=1552776240;
   	OWF_Key[86,6]:=51198609;
   	OWF_Key[86,7]:=746241045;
   	OWF_Key[86,8]:=229804881;
   	OWF_Key[87,0]:=1995108513;
   	OWF_Key[87,1]:=1307274145;
   	OWF_Key[87,2]:=1229662729;
   	OWF_Key[87,3]:=175094392;
   	OWF_Key[87,4]:=1994796318;
   	OWF_Key[87,5]:=1622102992;
   	OWF_Key[87,6]:=2105863629;
   	OWF_Key[87,7]:=1155246693;
   	OWF_Key[87,8]:=2139700852;
   	OWF_Key[88,0]:=1678496106;
   	OWF_Key[88,1]:=560336223;
   	OWF_Key[88,2]:=612456964;
   	OWF_Key[88,3]:=792857839;
   	OWF_Key[88,4]:=64320281;
   	OWF_Key[88,5]:=993892661;
   	OWF_Key[88,6]:=917072237;
   	OWF_Key[88,7]:=314456183;
   	OWF_Key[88,8]:=850885618;
   	OWF_Key[89,0]:=1027681791;
   	OWF_Key[89,1]:=548269312;
   	OWF_Key[89,2]:=599930273;
   	OWF_Key[89,3]:=835779663;
   	OWF_Key[89,4]:=12329049;
   	OWF_Key[89,5]:=2028885862;
   	OWF_Key[89,6]:=361691702;
   	OWF_Key[89,7]:=826916039;
   	OWF_Key[89,8]:=408464299;
   	OWF_Key[90,0]:=448193984;
   	OWF_Key[90,1]:=1587378053;
   	OWF_Key[90,2]:=888447072;
   	OWF_Key[90,3]:=1143626728;
   	OWF_Key[90,4]:=33082976;
   	OWF_Key[90,5]:=1341891390;
   	OWF_Key[90,6]:=1788734963;
   	OWF_Key[90,7]:=729549015;
   	OWF_Key[90,8]:=1847138909;
   	OWF_Key[91,0]:=463994107;
   	OWF_Key[91,1]:=102966428;
   	OWF_Key[91,2]:=873037777;
   	OWF_Key[91,3]:=617659960;
   	OWF_Key[91,4]:=522317748;
   	OWF_Key[91,5]:=935042477;
   	OWF_Key[91,6]:=1250501671;
   	OWF_Key[91,7]:=227117055;
   	OWF_Key[91,8]:=2061341368;
   	OWF_Key[92,0]:=1618315079;
   	OWF_Key[92,1]:=207922654;
   	OWF_Key[92,2]:=2075812444;
   	OWF_Key[92,3]:=121025035;
   	OWF_Key[92,4]:=1000281637;
   	OWF_Key[92,5]:=587174529;
   	OWF_Key[92,6]:=2053765231;
   	OWF_Key[92,7]:=2129245005;
   	OWF_Key[92,8]:=361288196;
   	OWF_Key[93,0]:=1353467296;
   	OWF_Key[93,1]:=501635479;
   	OWF_Key[93,2]:=485373383;
   	OWF_Key[93,3]:=939432416;
   	OWF_Key[93,4]:=775808151;
   	OWF_Key[93,5]:=1652196966;
   	OWF_Key[93,6]:=1122877217;
   	OWF_Key[93,7]:=2064732167;
   	OWF_Key[93,8]:=2045477847;
   	OWF_Key[94,0]:=1011797345;
   	OWF_Key[94,1]:=1066398681;
   	OWF_Key[94,2]:=230203801;
   	OWF_Key[94,3]:=348800200;
   	OWF_Key[94,4]:=1105596638;
   	OWF_Key[94,5]:=1315738884;
   	OWF_Key[94,6]:=1722507676;
   	OWF_Key[94,7]:=1134862033;
   	OWF_Key[94,8]:=1871676880;
   	OWF_Key[95,0]:=1425419837;
   	OWF_Key[95,1]:=275725913;
   	OWF_Key[95,2]:=1225884696;
   	OWF_Key[95,3]:=2028632425;
   	OWF_Key[95,4]:=1878874808;
   	OWF_Key[95,5]:=8711830;
   	OWF_Key[95,6]:=2091362778;
   	OWF_Key[95,7]:=472384707;
   	OWF_Key[95,8]:=1571264261;
   	OWF_Key[96,0]:=1902862333;
   	OWF_Key[96,1]:=728781155;
   	OWF_Key[96,2]:=948673298;
   	OWF_Key[96,3]:=1587481643;
   	OWF_Key[96,4]:=1323810487;
   	OWF_Key[96,5]:=736551736;
   	OWF_Key[96,6]:=1637521859;
   	OWF_Key[96,7]:=2020976519;
   	OWF_Key[96,8]:=1750183011;
   	OWF_Key[97,0]:=551889643;
   	OWF_Key[97,1]:=687738930;
   	OWF_Key[97,2]:=555893014;
   	OWF_Key[97,3]:=618811262;
   	OWF_Key[97,4]:=431374592;
   	OWF_Key[97,5]:=1543128027;
   	OWF_Key[97,6]:=2025661030;
   	OWF_Key[97,7]:=515207844;
   	OWF_Key[97,8]:=2034489760;
   	OWF_Key[98,0]:=1262881940;
   	OWF_Key[98,1]:=1393390823;
   	OWF_Key[98,2]:=508628527;
   	OWF_Key[98,3]:=1992308608;
   	OWF_Key[98,4]:=466953527;
   	OWF_Key[98,5]:=1077157707;
   	OWF_Key[98,6]:=742269167;
   	OWF_Key[98,7]:=1052679104;
   	OWF_Key[98,8]:=1453257683;
   	OWF_Key[99,0]:=379383308;
   	OWF_Key[99,1]:=72875063;
   	OWF_Key[99,2]:=1988889944;
   	OWF_Key[99,3]:=1371836394;
   	OWF_Key[99,4]:=1960344349;
   	OWF_Key[99,5]:=11428676;
   	OWF_Key[99,6]:=391563224;
   	OWF_Key[99,7]:=502976643;
   	OWF_Key[99,8]:=1931028225;
   	OWF_Key[100,0]:=1383341894;
   	OWF_Key[100,1]:=1427550471;
   	OWF_Key[100,2]:=1000912046;
   	OWF_Key[100,3]:=2018486416;
   	OWF_Key[100,4]:=1743274;
   	OWF_Key[100,5]:=2138437114;
   	OWF_Key[100,6]:=2004011284;
   	OWF_Key[100,7]:=1229119859;
   	OWF_Key[100,8]:=1852357095;
   	OWF_Key[101,0]:=1569957585;
   	OWF_Key[101,1]:=2118183153;
   	OWF_Key[101,2]:=1269113301;
   	OWF_Key[101,3]:=1852071747;
   	OWF_Key[101,4]:=1948776365;
   	OWF_Key[101,5]:=211752625;
   	OWF_Key[101,6]:=13134729;
   	OWF_Key[101,7]:=600508619;
   	OWF_Key[101,8]:=1035382672;
   	OWF_Key[102,0]:=2071585462;
   	OWF_Key[102,1]:=395724896;
   	OWF_Key[102,2]:=1017681513;
   	OWF_Key[102,3]:=1598707225;
   	OWF_Key[102,4]:=1359456368;
   	OWF_Key[102,5]:=1604516553;
   	OWF_Key[102,6]:=1673850999;
   	OWF_Key[102,7]:=1947342855;
   	OWF_Key[102,8]:=1331727978;
   	OWF_Key[103,0]:=3364383;
   	OWF_Key[103,1]:=280187649;
   	OWF_Key[103,2]:=970743292;
   	OWF_Key[103,3]:=168644725;
   	OWF_Key[103,4]:=1760852377;
   	OWF_Key[103,5]:=2021025184;
   	OWF_Key[103,6]:=1755513527;
   	OWF_Key[103,7]:=1238943457;
   	OWF_Key[103,8]:=1533747286;
   	OWF_Key[104,0]:=549107777;
   	OWF_Key[104,1]:=1242474044;
   	OWF_Key[104,2]:=439681614;
   	OWF_Key[104,3]:=945509569;
   	OWF_Key[104,4]:=1887607310;
   	OWF_Key[104,5]:=434280770;
   	OWF_Key[104,6]:=1397919920;
   	OWF_Key[104,7]:=1730690068;
   	OWF_Key[104,8]:=1756195635;
   	OWF_Key[105,0]:=985068248;
   	OWF_Key[105,1]:=1454164053;